// TIA Portal project "1215C_BREAKOUT_BOARD_IO-LINK_TEMPERATURE&TOWERLIGHT" (V19)

(* hardware
DEVICE "BREAKOUT_BOARD_PLC"  S7-1200 Station
   slot 0: "Rack_0"  S7-1200 Rack  Rack  V1.0
   slot 1: "BREAKOUT_BOARD_PLC"  CPU 1215C DC/DC/DC  6ES7 215-1AG40-0XB0  V4.6
DEVICE "BREAKOUT_BOARD_HMI"  KTP400 Basic PN
   slot 0: "BREAKOUT_BOARD_HMI"  KTP400 Basic PN  6AV2 123-2DB03-0AX0  16.0.0.0
   slot 1: "HMI_RT_1"  KTP400 Basic PN  6AV2 123-2DB03-0AX0  16.0.0.0
   slot 5: "BREAKOUT_BOARD_HMI.IE_CP_1"  PROFINET Interface  16.0.0.0
      slot 1: "PROFINET Interface"  PROFINET Interface
         slot 1: "Port_1"  Port
DEVICE "IFM_IO-LINK_MASTER"  GSD.Device.PN
   slot 0: "Rack"  Rack  V1.0
   slot 0: "AL1100"  AL1100  AL1100
      slot 0: "AL1100"  AL1100
      slot 1: "X1"  X1
         slot 1: "Port 1"  Port 1
         slot 2: "Port 2"  Port 2
      slot 1: "4 Ports_1"  4 Ports  AL1100
         slot 0: "IO-Link Master"  IO-Link Master
   slot 1: "IFM ITA2105 IO-Link In  2 Byte + PQI"  IO-Link In  2 Byte + PQI
   slot 2: "Banner TLF100 IO-Link Out 32 Byte + PQI"  IO-Link Out 32 Byte + PQI
   slot 3: "Disabled_P3"  Disabled
   slot 4: "Disabled_P4"  Disabled
DEVICE "SCALANCE XB008"  SCALANCE X-Station
   slot 0: "SCALANCE X rack"  Rail
   slot 0: "8PORT_SWITCH"  6GK5 008-0BA10-1AB2  V1.0
*)

// ===== PLC "BREAKOUT_BOARD_PLC"  CPU 1215C DC/DC/DC =====

VAR_GLOBAL   // PLC tag table "PLC_Outputs"
   "DQ0.0" AT %Q0.0 : Bool;   // Digital Output
   "DQ0.1" AT %Q0.1 : Bool;   // Digital Output
   "DQ0.2" AT %Q0.2 : Bool;   // Digital Output
   "DQ0.3" AT %Q0.3 : Bool;   // Digital Output
   "DQ0.4" AT %Q0.4 : Bool;   // Digital Output
   "DQ0.5" AT %Q0.5 : Bool;   // Digital Output
   "DQ0.6" AT %Q0.6 : Bool;   // Digital Output
   "DQ0.7" AT %Q0.7 : Bool;   // Digital Output
   "DQ1.0" AT %Q1.0 : Bool;   // Digital Output
   "DQ1.1" AT %Q1.1 : Bool;   // Digital Output
   "AQ0.0" AT %QW64 : Word;   // Analog Output
   "AQ0.1" AT %QW66 : Word;   // Analog Output
END_VAR

VAR_GLOBAL   // PLC tag table "PLC_Inputs"
   "DI0.0" AT %I0.0 : Bool;   // Digital Input
   "DI0.1" AT %I0.1 : Bool;   // Digital Input
   "DI0.2" AT %I0.2 : Bool;   // Digital Input
   "DI0.3" AT %I0.3 : Bool;   // Digital Input
   "DI0.4" AT %I0.4 : Bool;   // Digital Input
   "DI0.5" AT %I0.5 : Bool;   // Digital Input
   "DI0.6" AT %I0.6 : Bool;   // Digital Input
   "DI0.7" AT %I0.7 : Bool;   // Digital Input
   "DI1.0" AT %I1.0 : Bool;   // Digital Input
   "DI1.1" AT %I1.1 : Bool;   // Digital Input
   "DI1.2" AT %I1.2 : Bool;   // Digital Input
   "DI1.3" AT %I1.3 : Bool;   // Digital Input
   "DI1.4" AT %I1.4 : Bool;   // Digital Input
   "DI1.5" AT %I1.5 : Bool;   // Digital Input
   "AI0.0" AT %IW64 : Word;   // Analog Input
   "AI0.1" AT %IW66 : Word;   // Analog Input
END_VAR

VAR_GLOBAL   // PLC tag table "System_Tags"
   "Clock_Byte" AT %MB0 : Byte;
   "Clock_10Hz" AT %M0.0 : Bool;
   "Clock_5Hz" AT %M0.1 : Bool;
   "Clock_2.5Hz" AT %M0.2 : Bool;
   "Clock_2Hz" AT %M0.3 : Bool;
   "Clock_1.25Hz" AT %M0.4 : Bool;
   "Clock_1Hz" AT %M0.5 : Bool;
   "Clock_0.625Hz" AT %M0.6 : Bool;
   "Clock_0.5Hz" AT %M0.7 : Bool;
   "System_Byte" AT %MB1 : Byte;
   "FirstScan" AT %M1.0 : Bool;
   "DiagStatusUpdate" AT %M1.1 : Bool;
   "AlwaysTRUE" AT %M1.2 : Bool;
   "AlwaysFALSE" AT %M1.3 : Bool;
END_VAR

VAR_GLOBAL   // PLC tag table "Trigger_Tags"
   "xAQ_Trig" AT %M2.0 : Bool;
   "xTrig2" AT %M2.1 : Bool;
   "xTrig3" AT %M2.2 : Bool;
   "xTrig4" AT %M2.3 : Bool;
   "xTrig5" AT %M2.4 : Bool;
END_VAR

VAR_GLOBAL   // PLC tag table "IO-Link_Tags"
   "IFM_TA2105_Temp" AT %IW68 : Int;   // IO-Link Master X1
   "Banner_TLF100Pro_Byte0" AT %QB2 : Byte;   // IO-Link Master X2
   "Banner_TLF100Pro_Byte1" AT %QB3 : Byte;   // IO-Link Master X2
   "Banner_TLF100Pro_Byte2" AT %QB4 : Byte;   // IO-Link Master X2
   "Banner_TLF100Pro_Byte3" AT %QB5 : Byte;   // IO-Link Master X2
   "Banner_TLF100Pro_Byte4" AT %QB6 : Byte;   // IO-Link Master X2
   "Banner_TLF100Pro_Byte5" AT %QB7 : Byte;   // IO-Link Master X2
   "Banner_TLF100Pro_Byte6" AT %QB8 : Byte;   // IO-Link Master X2
   "Banner_TLF100Pro_Byte7" AT %QB9 : Byte;   // IO-Link Master X2
   "Banner_TLF100Pro_Byte8" AT %QB10 : Byte;   // IO-Link Master X2
   "Banner_TLF100Pro_Byte9" AT %QB11 : Byte;   // IO-Link Master X2
   "Banner_TLF100Pro_Byte10" AT %QB12 : Byte;   // IO-Link Master X2
   "Banner_TLF100Pro_Byte11" AT %QB13 : Byte;   // IO-Link Master X2
   "Banner_TLF100Pro_Byte12" AT %QB14 : Byte;   // IO-Link Master X2
   "Banner_TLF100Pro_Byte13" AT %QB15 : Byte;   // IO-Link Master X2
   "Banner_TLF100Pro_Byte14" AT %QB16 : Byte;   // IO-Link Master X2
   "Banner_TLF100Pro_Byte15" AT %QB17 : Byte;   // IO-Link Master X2
   "Banner_TLF100Pro_Byte16" AT %QB18 : Byte;   // IO-Link Master X2
   "Banner_TLF100Pro_Byte17" AT %QB19 : Byte;   // IO-Link Master X2
   "Banner_TLF100Pro_Byte18" AT %QB20 : Byte;   // IO-Link Master X2
   "Banner_TLF100Pro_Byte19" AT %QB21 : Byte;   // IO-Link Master X2
   "Banner_TLF100Pro_Byte20" AT %QB22 : Byte;   // IO-Link Master X2
   "Banner_TLF100Pro_Byte21" AT %QB23 : Byte;   // IO-Link Master X2
   "Banner_TLF100Pro_Byte22" AT %QB24 : Byte;   // IO-Link Master X2 - Not Used
   "Banner_TLF100Pro_Byte23" AT %QB25 : Byte;   // IO-Link Master X2 - Not Used
   "Banner_TLF100Pro_Byte24" AT %QB26 : Byte;   // IO-Link Master X2 - Not Used
   "Banner_TLF100Pro_Byte25" AT %QB27 : Byte;   // IO-Link Master X2 - Not Used
   "Banner_TLF100Pro_Byte26" AT %QB28 : Byte;   // IO-Link Master X2 - Not Used
   "Banner_TLF100Pro_Byte27" AT %QB29 : Byte;   // IO-Link Master X2 - Not Used
   "Banner_TLF100Pro_Byte28" AT %QB30 : Byte;   // IO-Link Master X2 - Not Used
   "Banner_TLF100Pro_Byte29" AT %QB31 : Byte;   // IO-Link Master X2 - Not Used
   "Banner_TLF100Pro_Byte30" AT %QB32 : Byte;   // IO-Link Master X2 - Not Used
   "Banner_TLF100Pro_Byte31" AT %QB33 : Byte;   // IO-Link Master X2 - Not Used
END_VAR

// folder: WS01_TVET_Workstation/00-I/O_Mapping

DATA_BLOCK "DB001-PLC_I/O"   // DB1
TITLE = PLC I/O Global Database
{ S7_Optimized_Access := 'TRUE' }
VERSION : 0.1
// Variables used to mirror the physical PLC I/O states.
   VAR
      Inputs : Struct   // PLC Inputs Structure
         "xDI0.0" : Bool;
         "xDI0.1" : Bool;
         "xDI0.2" : Bool;
         "xDI0.3" : Bool;
         "xDI0.4" : Bool;
         "xDI0.5" : Bool;
         "xDI0.6" : Bool;
         "xDI0.7" : Bool;
         "xDI1.0" : Bool;
         "xDI1.1" : Bool;
         "xDI1.2" : Bool;
         "xDI1.3" : Bool;
         "xDI1.4" : Bool;
         "xDI1.5" : Bool;
         "rAI0.0_Scaled" : Real;   // 0 to 24648 = 0 to 10 V
         "rAI0.1_Scaled" : Real;   // 0 to 24648 = 0 to 10 V
      END_STRUCT;
      Outputs : Struct   // PLC Outputs Structure
         "xDQ0.0" : Bool;
         "xDQ0.1" : Bool;
         "xDQ0.2" : Bool;
         "xDQ0.3" : Bool;
         "xDQ0.4" : Bool;
         "xDQ0.5" : Bool;
         "xDQ0.6" : Bool;
         "xDQ0.7" : Bool;
         "xDQ1.0" : Bool;
         "xDQ1.1" : Bool;
         "iAQ0.0_RAW" : Int := 0;
         "rAQ0.0_Scaled" : Real;   // 0 to 24648 = 0 to 20 mA
         "iAQ0.1_RAW" : Int := 0;
         "rAQ0.1_Scaled" : Real;   // 0 to 24648 = 0 to 20 mA
      END_STRUCT;
   END_VAR
BEGIN
END_DATA_BLOCK

DATA_BLOCK "DB003-IO-Link_I/O"   // DB3
TITLE = IO-Link I/O Global Database
{ S7_Optimized_Access := 'TRUE' }
VERSION : 0.1
// Variables used to mirror the physical IO-Link I/O states.
   VAR
      Inputs : Struct   // IO-Link Inputs Structure
         wTemp_RAW : Word;   // Temperature Sensor Scaled Value
      END_STRUCT;
      Outputs : Struct   // IO-Link Outputs Structure
         TL_Byte_Array : Array[0..21] of Byte;   // Tower Light Byte Array
      END_STRUCT;
   END_VAR
BEGIN
END_DATA_BLOCK

// folder: WS01_TVET_Workstation/01-DateTime

DATA_BLOCK "DB002-DateTime"   // DB2
TITLE = PLC Date/Time Global Database
{ S7_Optimized_Access := 'TRUE' }
VERSION : 0.1
// Variables used to store the PLC date/time & custom date/time formatting.
   VAR
      RD_LOC_T_Ret : Int := 0;   // Return value for Read Local Time Block
      LOCAL_DTL : DTL := DTL#1970-01-01-00:00:00;   // RAW DTL
      "Date" : Date := D#1990-01-01;   // RAW Date
      "Time" : Time_Of_Day := TOD#00:00:00;   // RAW Time
      DTLtoString_Ret : String;   // Return value for DTL to String Block
      sCustomDate_YY : String := '';   // Custom year
      sCustomDate_MM : String := '';   // Custom month
      sCustomDate_DD : String := '';   // Custom Day
      sCustomTime_HH : String := '';   // Custom hour
      sCustomTime_MM : String := '';   // Custom minute
      sCustomDate_DDMMYY : String := '';   // Custom date format
      sCustomTime_HHMM : String := '';   // Custom time format
   END_VAR
BEGIN
END_DATA_BLOCK

// folder: WS01_TVET_Workstation/02-IOLink_Control

DATA_BLOCK "DB003-IOLink_Data"   // DB4
TITLE = IO-Link Data Global Database
{ S7_Optimized_Access := 'TRUE' }
VERSION : 0.1
// Variables used to process data from connected devices.
   VAR
      TempSensor_Data : Struct   // Temperature Sensor Data Structure
         rDeg_C : Real;   // Degrees Celsius
         rDeg_F : Real;   // Degrees Fahrenheit
      END_STRUCT;
      TL_ProcessData : Struct   // Tower Light Process Data Structure
         Animations : Struct   // Animation Parameters Structure
            iOff : Int := 0;   // Animations
            iSteady : Int := 1;   // Animations
            iFlash : Int := 2;   // Animations
            i2ColourFlash : Int := 3;   // Animations
            i2ColourShift : Int := 4;   // Animations
            iEndsSteady : Int := 5;   // Animations
            iEndsFlash : Int := 6;   // Animations
            iScroll : Int := 7;   // Animations
            iCenterScroll : Int := 8;   // Animations
            iBounce : Int := 9;   // Animations
            iCenterBounce : Int := 10;   // Animations
            iIntensitySweep : Int := 11;   // Animations
            i2ColourSweep : Int := 12;   // Animations
            iSpectrum : Int := 13;   // Animations
            iLevelSteady : Int := 14;   // Animations
            iLevelFlash : Int := 15;   // Animations
         END_STRUCT;
         Colours : Struct   // Colour Parameters Structure
            iGreen : Int := 0;   // Colours
            iRed : Int := 1;   // Colours
            iOrange : Int := 2;   // Colours
            iAmber : Int := 3;   // Colours
            iYellow : Int := 4;   // Colours
            iLimeGreen : Int := 5;   // Colours
            iSpringGreen : Int := 6;   // Colours
            iCyan : Int := 7;   // Colours
            iSkyBlue : Int := 8;   // Colours
            iBlue : Int := 9;   // Colours
            iViolet : Int := 10;   // Colours
            iMegenta : Int := 11;   // Colours
            iRose : Int := 12;   // Colours
            iDaylightWhite : Int := 13;   // Colours
         END_STRUCT;
         ColourIntensities : Struct   // Colour Intensity Parameters Structure
            iHigh : Int := 0;   // Colour Intensity
            iLow : Int := 1;   // Colour Intensity
            iMedium : Int := 2;   // Colour Intensity
            iOff : Int := 3;   // Colour Intensity
         END_STRUCT;
         Speeds : Struct   // Speed Parameters Structure
            iMedium : Int := 0;   // Speed
            iFast : Int := 1;   // Speed
            iSlow : Int := 2;   // Speed
         END_STRUCT;
         PulsePatterns : Struct   // Pulse Pattern Parameters Structure
            iNormal : Int := 0;   // Pulse Pattern
            iStrobe : Int := 1;   // Pulse Pattern
            i3Pulse : Int := 2;   // Pulse Pattern
            iSOS : Int := 3;   // Pulse Pattern
            iRandom : Int := 4;   // Pulse Pattern
         END_STRUCT;
         ScrollStyles : Struct   // Scroll Style Parameters Structure
            iSolid : Int := 0;   // Scroll Style
            iTail : Int := 1;   // Scroll Style
            iRipple : Int := 2;   // Scroll Style
         END_STRUCT;
         Directions : Struct   // Direction Parameters Structure
            xUp : Bool := FALSE;   // Direction
            xDown : Bool := TRUE;   // Direction
         END_STRUCT;
         iColourWidthPercent : Int := 100;   // Percent Width of Colour (1-100)
         AudibleTypes : Struct   // Audible Type Parameters Structure
            iPulse : Int := 0;   // Audible Type
            iWobble : Int := 1;   // Audible Type
            iStrobe : Int := 2;   // Audible Type
            iWhoop : Int := 4;   // Audible Type
            iStaccato : Int := 5;   // Audible Type
            iSiren : Int := 6;   // Audible Type
            iContinuous1 : Int := 8;   // Audible Type
            iContinuous2 : Int := 9;   // Audible Type
            iJungle : Int := 16;   // Audible Type
            iMelody1 : Int := 17;   // Audible Type
            iMelody2 : Int := 18;   // Audible Type
            iMelody3 : Int := 19;   // Audible Type
         END_STRUCT;
         AudibleVolumes : Struct   // Audible Volume Parameters Structure
            iOff : Int := 0;   // Audible Volume
            iLow : Int := 1;   // Audible Volume
            iMedium : Int := 2;   // Audible Volume
            iHigh : Int := 3;   // Audible Volume
         END_STRUCT;
      END_STRUCT;
   END_VAR
BEGIN
END_DATA_BLOCK

// folder: WS01_TVET_Workstation/03-HMI_Control

DATA_BLOCK "DB005-HMI_Data"   // DB5
TITLE = HMI Data Global Database
{ S7_Optimized_Access := 'TRUE' }
VERSION : 0.1
// Variables used to process data from the HMI.
   VAR
      iScreen_Number : UInt;   // HMI Active Screen Number
      TowerLight : Struct   // Tower Light HMI Variables Structure
         Segment1 : Struct   // Segment 1 Structure
            iAnimate : Int;   // Animations
            iSavedAnimate : Int;   // Saved Animation Value
            iColour1 : Int;   // Colour1 Colours
            iColour2 : Int;   // Colour2 Colours
            iSpeed : Int;   // Speeds
            "iClrWidth%" : Int := 100;   // Colour Width Percentage
         END_STRUCT;
         Segment2 : Struct   // Segment 2 Structure
            iAnimate : Int;   // Animations
            iSavedAnimate : Int;   // Saved Animation Value
            iColour1 : Int;   // Colour1 Colours
            iColour2 : Int;   // Colour2 Colours
            iSpeed : Int;   // Speeds
            "iClrWidth%" : Int := 100;   // Colour Width Percentage
         END_STRUCT;
         Segment3 : Struct   // Segment 3 Structure
            iAnimate : Int;   // Animations
            iSavedAnimate : Int;   // Saved Animation Value
            iColour1 : Int;   // Colour1 Colours
            iColour2 : Int;   // Colour2 Colours
            iSpeed : Int;   // Speeds
            "iClrWidth%" : Int := 100;   // Colour Width Percentage
         END_STRUCT;
         Audible : Struct   // Audible (Sound) Structure
            iType : Int;   // Types
            iVolume : Int;   // Volumes
            iSavedVolume : Int;   // Saved Volume Value
         END_STRUCT;
         xSave_Config : Bool;   // Save Tower Light Configs Button
      END_STRUCT;
   END_VAR
BEGIN
END_DATA_BLOCK

// folder: (top level)

ORGANIZATION_BLOCK "Main"   // OB1, LAD, ProgramCycle
TITLE = "Main Program Sweep (Cycle)"
{ S7_Optimized_Access := 'TRUE' }
VERSION : 0.1
   VAR_INPUT
      Initial_Call : Bool;   // Initial call of this OB
      Remanence : Bool;   // =True, if remanent data are available
   END_VAR
BEGIN

REGION Network 1 (SCL): ================= PROGRAM_INFORMATION =================
   (*
   ==================================================================
   ********************* PLC I/O BREAKOUT BOARD *********************
   ==================================================================

   TVET Workstation WS01:
   1215C DC/DC/DC - 6ES7215-1AG40-0XB0 - IP: 192.168.0.175/24

   KTP400 HMI - 6AV2123-2DB03-0AX0 - IP: 192.168.0.176/24

   IFM IO-Link Master - AL1100 - IP: 192.168.0.177/24

   =======================================================================

   The program has 4 main sections:
   - Date/Time Handler,
   - I/O Handlers,
   - IO-Link Devices Handler,
   - HMI Handler.

   Date/Time Handler FC:
   - local PLC date/time is read & formatted into a 24HR time & DD/MM/YYYY.

   I/O Handler FCs:
   - maps the physical PLC inputs & outputs to corresponding tags in DB001,
   - handles scaling of the PLC Analog I/O,
   - maps the IO-Link inputs & outputs to corresponding tags in DB003,
   - ensures that physical I/O tags are only used once in the code.

   IO-Link Device Handler FCs:
   - connected IO-Link devices are controlled in this section:
       - the temperature sensor conversion logic is handled by an IFM
         provided FC which scales the input value & converts to Fahrenheit.
       - the tower light ON/OFF logic is handled by the TowerLight Handler FC.
   - create & call new FC's for any additional IO-Link devices that may
     get added.

   Additional Notes:
   PLC Tags grouped according to their use/function.

   =======================================================================

   Analog Input Technical data:
   - Number of inputs: 2
   - Type: Voltage (single-ended)
   - Full-scale range: 0 to 10 V
   - Full-scale range (data word): 0 to 27648
   - Overshoot range: 10.001 to 11.759 V
   - Overshoot range (data word): 27649 to 32511
   - Overflow range: 11.760 to 11.852 V
   - Overflow range (data word): 32512 to 32767
   - Resolution: 10 bits
   - Maximum withstand voltage: 35 V DC
   - Smoothing: None, Weak, Medium, or Strong
   - Noise rejection: 10, 50, or 60 Hz
   - Impedance: ≥100 KΩ
   - Isolation (field side to logic): None
   - Accuracy (25 °C / -20 to 60 °C): 3.0% / 3.5% of full-scale
   - Cable length (meters): 100 m, shielded twisted pair
   - Rated range: 0     = 0 V
                  34    = 12 mV
                  20736 = 7.5 V
                  27648 = 10 V

   =======================================================================

   Analog Output Technical data:
   - Number of outputs: 2
   - Type: Current
   - Full-scale range: 0 to 20 mA
   - Full-scale range (data word): 0 to 27648
   - Overshoot range: 20.01 to 23.52 mA
   - Overshoot range (data word): 27649 to 32511
   - Overflow range data word: 32512 to 32767
   - Resolution: 10 bits
   - Output drive impedance: ≤500 Ω max
   - Isolation (field side to logic): None
   - Accuracy (25 °C / -20 to 60 °C): 3.0% / 3.5% of full-scale
   - Settling time: 2 ms
   - Cable length (meters): 100 m, shielded twisted pair
   - Rated range: 0     = 0 mA
                  34    = 0.0247 mA
                  20736 = 15 mA
                  27648 = 20 mA

   =======================================================================

   TA2105 IO-Link Temperature Transmitter documentation:
   https://www.ifm.com/us/en/product/TA2105#documents

   Process Data In length = 2bytes

   The IO-Link Inputs screen on the HMI displays a bar graph of the current
   measured temperature for the sensor connected to port X1.

   =======================================================================

   TLF100Pro IO-Link Tower Light Data Reference Guide:
   www.bannerengineering.com/us/en/products/part.812293.html

   Process Data Out length = 22bytes

   Modes:
   - Segment Mode
   - Run Mode
   - Advanced Mode
   - Level Mode

   We will be using the "Advanced Mode" to configure Segments 1, 2, 3
   and Audible. Segment 4 can be ignored as it is not applicable to
   this tower light model.

   The function interface contains a list of the available parameters
   that can be used to set segment bytes.

   Each colour segment has 5 bytes that need to be set with a
   corresponding constant value to configure the segment.

   The audible (segment) has 2 bytes that need to be set with a
   corresponding constant value.

   Segment bytes are defined as follows:
   -----------------------------
   > Segement 1 - byte 21 to 17:
       - 21 = Animation (8bits)
       - 20 = Colour1 (5bits) + Intensity (3bits)
       - 19 = Colour2 (5bits) + Intensity (3bits)
       - 18 = Speed (2bits) + Pulse Pattern (3bits) + Style (2bits) + Direction (1bit)
       - 17 = Colour Width Percentage (1-100)
   -----------------------------
   > Segement 2 - byte 16 to 12:
       - 16 = Animation (8bits)
       - 15 = Colour1 (5bits) + Intensity (3bits)
       - 14 = Colour2 (5bits) + Intensity (3bits)
       - 13 = Speed (2bits) + Pulse Pattern (3bits) + Style (2bits) + Direction (1bit)
       - 12 = Colour Width Percentage (1-100)
   ----------------------------
   > Segement 3 - byte 11 to 7:
       - 11 = Animation (8bits)
       - 10 = Colour1 (5bits) + Intensity (3bits)
       - 09 = Colour2 (5bits) + Intensity (3bits)
       - 08 = Speed (2bits) + Pulse Pattern (3bits) + Style (2bits) + Direction (1bit)
       - 07 = Colour Width Percentage (1-100)
   ---------------------------
   > Segement 4 - byte 6 to 2: !!NOT USED!!
       - 06 = Animation (8bits)
       - 05 = Colour1 (5bits) + Intensity (3bits)
       - 04 = Colour2 (5bits) + Intensity (3bits)
       - 03 = Speed (2bits) + Pulse Pattern (3bits) + Style (2bits) + Direction (1bit)
       - 02 = Colour Width Percentage (1-100)
   ------------------------
   > Audible - byte 1 to 0:
       - 01 = Type (8bits)
       - 00 = Volume (8bits)

   Some segment bytes are divided into sub-indexes depending on the 
   functions available for a particular byte.

   Since we are aiming at creating basic functionality
   (basic solid or flashing colours & sound)
   we will ignore many of the sub-indexes functions & simply set the
   entire byte with a single parameter constant.

   Segment parameters are set via the HMI and controlled via input
   switches.

   =======================================================================
   *)
END_REGION

REGION Network 2: ================= LOCAL_DATE/TIME =================
END_REGION

REGION Network 3: Call the Date/Time Handler Function
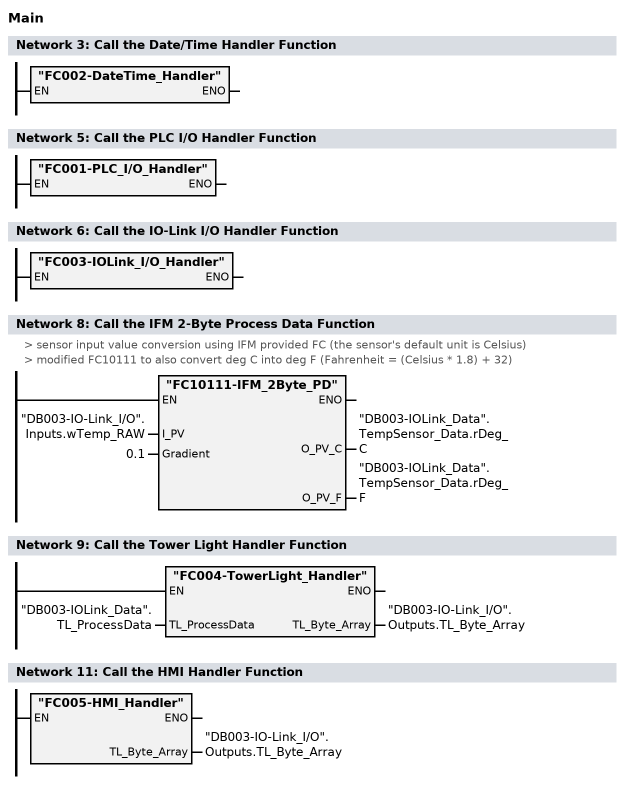
   RUNG wire#powerrail
      "FC002-DateTime_Handler"()
   END_RUNG
   // the same network as SCL:
   "FC002-DateTime_Handler"();
END_REGION

REGION Network 4: ================= I/O_MAPPING =================
END_REGION

REGION Network 5: Call the PLC I/O Handler Function
   RUNG wire#powerrail
      "FC001-PLC_I/O_Handler"()
   END_RUNG
   // the same network as SCL:
   "FC001-PLC_I/O_Handler"();
END_REGION

REGION Network 6: Call the IO-Link I/O Handler Function
   RUNG wire#powerrail
      "FC003-IOLink_I/O_Handler"()
   END_RUNG
   // the same network as SCL:
   "FC003-IOLink_I/O_Handler"();
END_REGION

REGION Network 7: ================= IO-LINK_DEVICES =================
END_REGION

REGION Network 8: Call the IFM 2-Byte Process Data Function
   // > sensor input value conversion using IFM provided FC (the sensor's default unit is Celsius)
   // > modified FC10111 to also convert deg C into deg F (Fahrenheit = (Celsius * 1.8) + 32)
   RUNG wire#powerrail
      "FC10111-IFM_2Byte_PD"(I_PV := "DB003-IO-Link_I/O".Inputs.wTemp_RAW, Gradient := 0.1, O_PV_C => "DB003-IOLink_Data".TempSensor_Data.rDeg_C, O_PV_F => "DB003-IOLink_Data".TempSensor_Data.rDeg_F)
   END_RUNG
   // the same network as SCL:
   "FC10111-IFM_2Byte_PD"(I_PV := "DB003-IO-Link_I/O".Inputs.wTemp_RAW,
                          Gradient := 0.1,
                          O_PV_C => "DB003-IOLink_Data".TempSensor_Data.rDeg_C,
                          O_PV_F => "DB003-IOLink_Data".TempSensor_Data.rDeg_F);
END_REGION

REGION Network 9: Call the Tower Light Handler Function
   RUNG wire#powerrail
      "FC004-TowerLight_Handler"(TL_ProcessData := "DB003-IOLink_Data".TL_ProcessData, TL_Byte_Array => "DB003-IO-Link_I/O".Outputs.TL_Byte_Array)
   END_RUNG
   // the same network as SCL:
   "FC004-TowerLight_Handler"(TL_ProcessData := "DB003-IOLink_Data".TL_ProcessData,
                           TL_Byte_Array => "DB003-IO-Link_I/O".Outputs.TL_Byte_Array);
END_REGION

REGION Network 10: ================= HMI_CONTROL =================
END_REGION

REGION Network 11: Call the HMI Handler Function
   RUNG wire#powerrail
      "FC005-HMI_Handler"(TL_Byte_Array => "DB003-IO-Link_I/O".Outputs.TL_Byte_Array)
   END_RUNG
   // the same network as SCL:
   "FC005-HMI_Handler"(TL_Byte_Array => "DB003-IO-Link_I/O".Outputs.TL_Byte_Array);
END_REGION
END_ORGANIZATION_BLOCK

// folder: WS01_TVET_Workstation/00-I/O_Mapping

FUNCTION "FC001-PLC_I/O_Handler" : Void   // FC1, LAD
TITLE = PLC Input Output Handler
{ S7_Optimized_Access := 'TRUE' }
VERSION : 0.1
// This function block is for interfacing the physical PLC input/output connections to a Global DB's (DB001-PLC_I/O for ).
   VAR_TEMP
      "rAI0.0_Temp" : Real;
      "rAI0.1_Temp" : Real;
      "rAQ0.0_Temp" : Real;
      "rAQ0.1_Temp" : Real;
   END_VAR
   VAR_TEMP   // added for the SCL form of the ladder/FBD networks
      _w1 : Bool;
   END_VAR
BEGIN

REGION Network 1: ================= DIGITAL_INPUTS =================
END_REGION

REGION Network 2: BANK_0
   // > DI0.0 - DI0.7
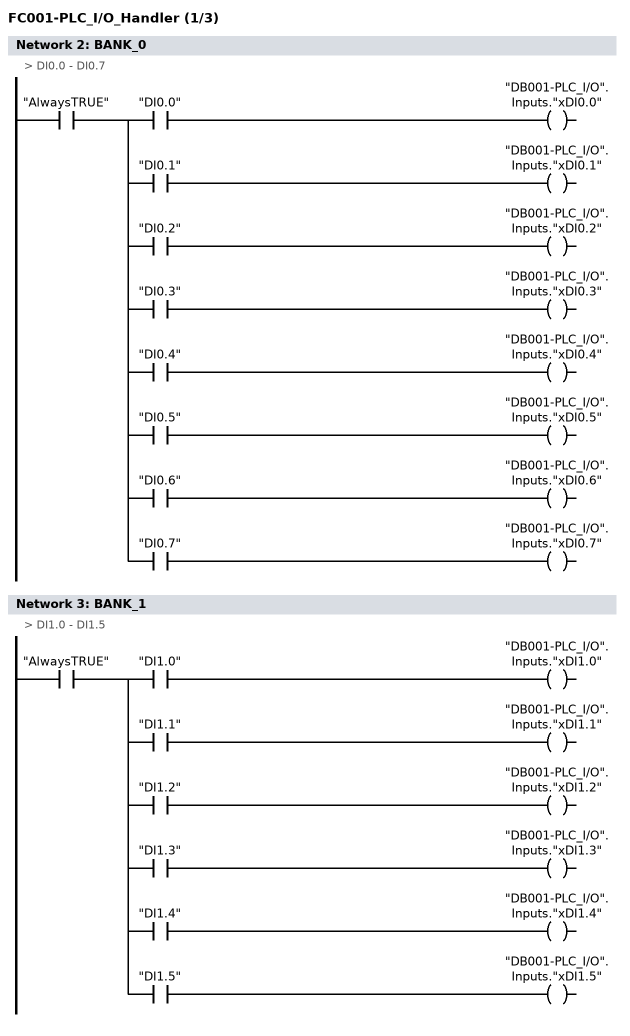
   RUNG wire#powerrail
      Contact( "AlwaysTRUE" )
      wire#w1
      Contact( "DI0.0" )
      Coil( "DB001-PLC_I/O".Inputs."xDI0.0" )
   END_RUNG
   RUNG wire#w1
      Contact( "DI0.1" )
      Coil( "DB001-PLC_I/O".Inputs."xDI0.1" )
   END_RUNG
   RUNG wire#w1
      Contact( "DI0.2" )
      Coil( "DB001-PLC_I/O".Inputs."xDI0.2" )
   END_RUNG
   RUNG wire#w1
      Contact( "DI0.3" )
      Coil( "DB001-PLC_I/O".Inputs."xDI0.3" )
   END_RUNG
   RUNG wire#w1
      Contact( "DI0.4" )
      Coil( "DB001-PLC_I/O".Inputs."xDI0.4" )
   END_RUNG
   RUNG wire#w1
      Contact( "DI0.5" )
      Coil( "DB001-PLC_I/O".Inputs."xDI0.5" )
   END_RUNG
   RUNG wire#w1
      Contact( "DI0.6" )
      Coil( "DB001-PLC_I/O".Inputs."xDI0.6" )
   END_RUNG
   RUNG wire#w1
      Contact( "DI0.7" )
      Coil( "DB001-PLC_I/O".Inputs."xDI0.7" )
   END_RUNG
   // the same network as SCL:
   "DB001-PLC_I/O".Inputs."xDI0.0" := "AlwaysTRUE" AND "DI0.0";
   "DB001-PLC_I/O".Inputs."xDI0.1" := "AlwaysTRUE" AND "DI0.1";
   "DB001-PLC_I/O".Inputs."xDI0.2" := "AlwaysTRUE" AND "DI0.2";
   "DB001-PLC_I/O".Inputs."xDI0.3" := "AlwaysTRUE" AND "DI0.3";
   "DB001-PLC_I/O".Inputs."xDI0.4" := "AlwaysTRUE" AND "DI0.4";
   "DB001-PLC_I/O".Inputs."xDI0.5" := "AlwaysTRUE" AND "DI0.5";
   "DB001-PLC_I/O".Inputs."xDI0.6" := "AlwaysTRUE" AND "DI0.6";
   "DB001-PLC_I/O".Inputs."xDI0.7" := "AlwaysTRUE" AND "DI0.7";
END_REGION

REGION Network 3: BANK_1
   // > DI1.0 - DI1.5
   RUNG wire#powerrail
      Contact( "AlwaysTRUE" )
      wire#w1
      Contact( "DI1.0" )
      Coil( "DB001-PLC_I/O".Inputs."xDI1.0" )
   END_RUNG
   RUNG wire#w1
      Contact( "DI1.1" )
      Coil( "DB001-PLC_I/O".Inputs."xDI1.1" )
   END_RUNG
   RUNG wire#w1
      Contact( "DI1.2" )
      Coil( "DB001-PLC_I/O".Inputs."xDI1.2" )
   END_RUNG
   RUNG wire#w1
      Contact( "DI1.3" )
      Coil( "DB001-PLC_I/O".Inputs."xDI1.3" )
   END_RUNG
   RUNG wire#w1
      Contact( "DI1.4" )
      Coil( "DB001-PLC_I/O".Inputs."xDI1.4" )
   END_RUNG
   RUNG wire#w1
      Contact( "DI1.5" )
      Coil( "DB001-PLC_I/O".Inputs."xDI1.5" )
   END_RUNG
   // the same network as SCL:
   "DB001-PLC_I/O".Inputs."xDI1.0" := "AlwaysTRUE" AND "DI1.0";
   "DB001-PLC_I/O".Inputs."xDI1.1" := "AlwaysTRUE" AND "DI1.1";
   "DB001-PLC_I/O".Inputs."xDI1.2" := "AlwaysTRUE" AND "DI1.2";
   "DB001-PLC_I/O".Inputs."xDI1.3" := "AlwaysTRUE" AND "DI1.3";
   "DB001-PLC_I/O".Inputs."xDI1.4" := "AlwaysTRUE" AND "DI1.4";
   "DB001-PLC_I/O".Inputs."xDI1.5" := "AlwaysTRUE" AND "DI1.5";
END_REGION

REGION Network 4: ================= DIGITAL_OUTPUTS =================
END_REGION

REGION Network 5: BANK_0
   // > DQ0.0 - DQ0.7
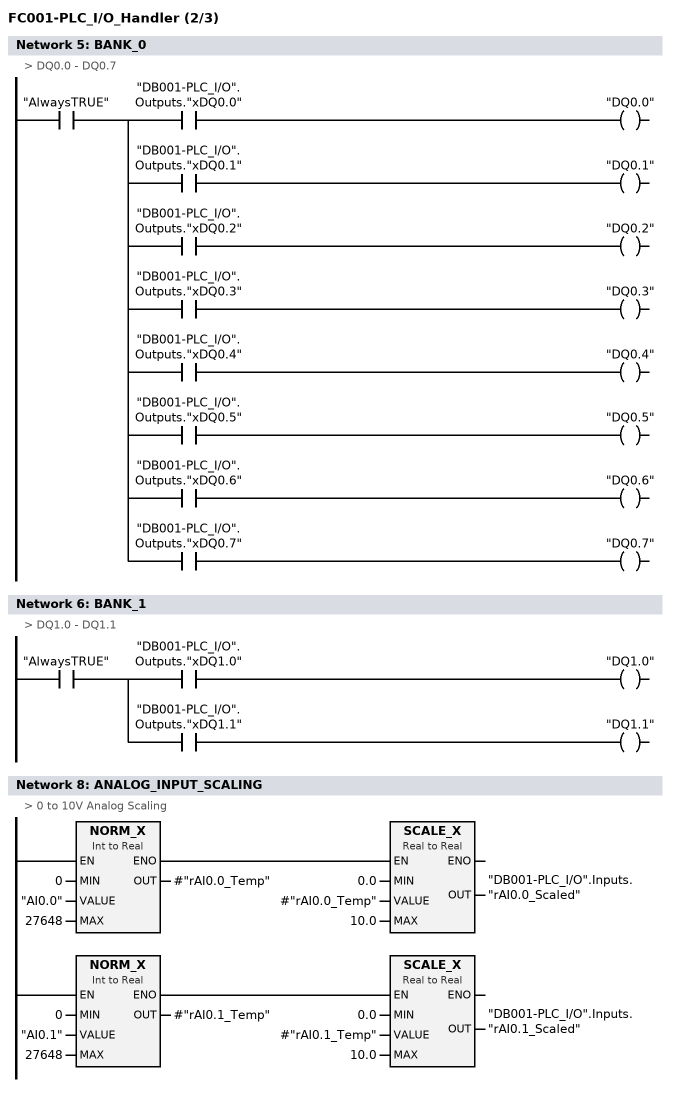
   RUNG wire#powerrail
      Contact( "AlwaysTRUE" )
      wire#w1
      Contact( "DB001-PLC_I/O".Outputs."xDQ0.0" )
      Coil( "DQ0.0" )
   END_RUNG
   RUNG wire#w1
      Contact( "DB001-PLC_I/O".Outputs."xDQ0.1" )
      Coil( "DQ0.1" )
   END_RUNG
   RUNG wire#w1
      Contact( "DB001-PLC_I/O".Outputs."xDQ0.2" )
      Coil( "DQ0.2" )
   END_RUNG
   RUNG wire#w1
      Contact( "DB001-PLC_I/O".Outputs."xDQ0.3" )
      Coil( "DQ0.3" )
   END_RUNG
   RUNG wire#w1
      Contact( "DB001-PLC_I/O".Outputs."xDQ0.4" )
      Coil( "DQ0.4" )
   END_RUNG
   RUNG wire#w1
      Contact( "DB001-PLC_I/O".Outputs."xDQ0.5" )
      Coil( "DQ0.5" )
   END_RUNG
   RUNG wire#w1
      Contact( "DB001-PLC_I/O".Outputs."xDQ0.6" )
      Coil( "DQ0.6" )
   END_RUNG
   RUNG wire#w1
      Contact( "DB001-PLC_I/O".Outputs."xDQ0.7" )
      Coil( "DQ0.7" )
   END_RUNG
   // the same network as SCL:
   "DQ0.0" := "AlwaysTRUE" AND "DB001-PLC_I/O".Outputs."xDQ0.0";
   "DQ0.1" := "AlwaysTRUE" AND "DB001-PLC_I/O".Outputs."xDQ0.1";
   "DQ0.2" := "AlwaysTRUE" AND "DB001-PLC_I/O".Outputs."xDQ0.2";
   "DQ0.3" := "AlwaysTRUE" AND "DB001-PLC_I/O".Outputs."xDQ0.3";
   "DQ0.4" := "AlwaysTRUE" AND "DB001-PLC_I/O".Outputs."xDQ0.4";
   "DQ0.5" := "AlwaysTRUE" AND "DB001-PLC_I/O".Outputs."xDQ0.5";
   "DQ0.6" := "AlwaysTRUE" AND "DB001-PLC_I/O".Outputs."xDQ0.6";
   "DQ0.7" := "AlwaysTRUE" AND "DB001-PLC_I/O".Outputs."xDQ0.7";
END_REGION

REGION Network 6: BANK_1
   // > DQ1.0 - DQ1.1
   RUNG wire#powerrail
      Contact( "AlwaysTRUE" )
      wire#w1
      Contact( "DB001-PLC_I/O".Outputs."xDQ1.0" )
      Coil( "DQ1.0" )
   END_RUNG
   RUNG wire#w1
      Contact( "DB001-PLC_I/O".Outputs."xDQ1.1" )
      Coil( "DQ1.1" )
   END_RUNG
   // the same network as SCL:
   "DQ1.0" := "AlwaysTRUE" AND "DB001-PLC_I/O".Outputs."xDQ1.0";
   "DQ1.1" := "AlwaysTRUE" AND "DB001-PLC_I/O".Outputs."xDQ1.1";
END_REGION

REGION Network 7: ================= ANALOG_PROCESSING =================
END_REGION

REGION Network 8: ANALOG_INPUT_SCALING
   // > 0 to 10V Analog Scaling
   RUNG wire#powerrail
      { S7_Templates := "[SrcType := Int, DestType := Real]" } Normalize(min := 0, value := "AI0.0", max := 27648, out => #"rAI0.0_Temp")
      { S7_Templates := "[SrcType := Real, DestType := Real]" } Scale(min := 0.0, value := #"rAI0.0_Temp", max := 10.0, out => "DB001-PLC_I/O".Inputs."rAI0.0_Scaled")
   END_RUNG
   RUNG wire#powerrail
      { S7_Templates := "[SrcType := Int, DestType := Real]" } Normalize(min := 0, value := "AI0.1", max := 27648, out => #"rAI0.1_Temp")
      { S7_Templates := "[SrcType := Real, DestType := Real]" } Scale(min := 0.0, value := #"rAI0.1_Temp", max := 10.0, out => "DB001-PLC_I/O".Inputs."rAI0.1_Scaled")
   END_RUNG
   // the same network as SCL:
   #"rAI0.0_Temp" := NORM_X(MIN := 0, VALUE := "AI0.0", MAX := 27648);
   "DB001-PLC_I/O".Inputs."rAI0.0_Scaled" := SCALE_X(MIN := 0.0, VALUE := #"rAI0.0_Temp", MAX := 10.0);
   #"rAI0.1_Temp" := NORM_X(MIN := 0, VALUE := "AI0.1", MAX := 27648);
   "DB001-PLC_I/O".Inputs."rAI0.1_Scaled" := SCALE_X(MIN := 0.0, VALUE := #"rAI0.1_Temp", MAX := 10.0);
END_REGION

REGION Network 9: ANALOG_OUTPUT_SCALING
   // > 0 to 20mA Analog Scaling
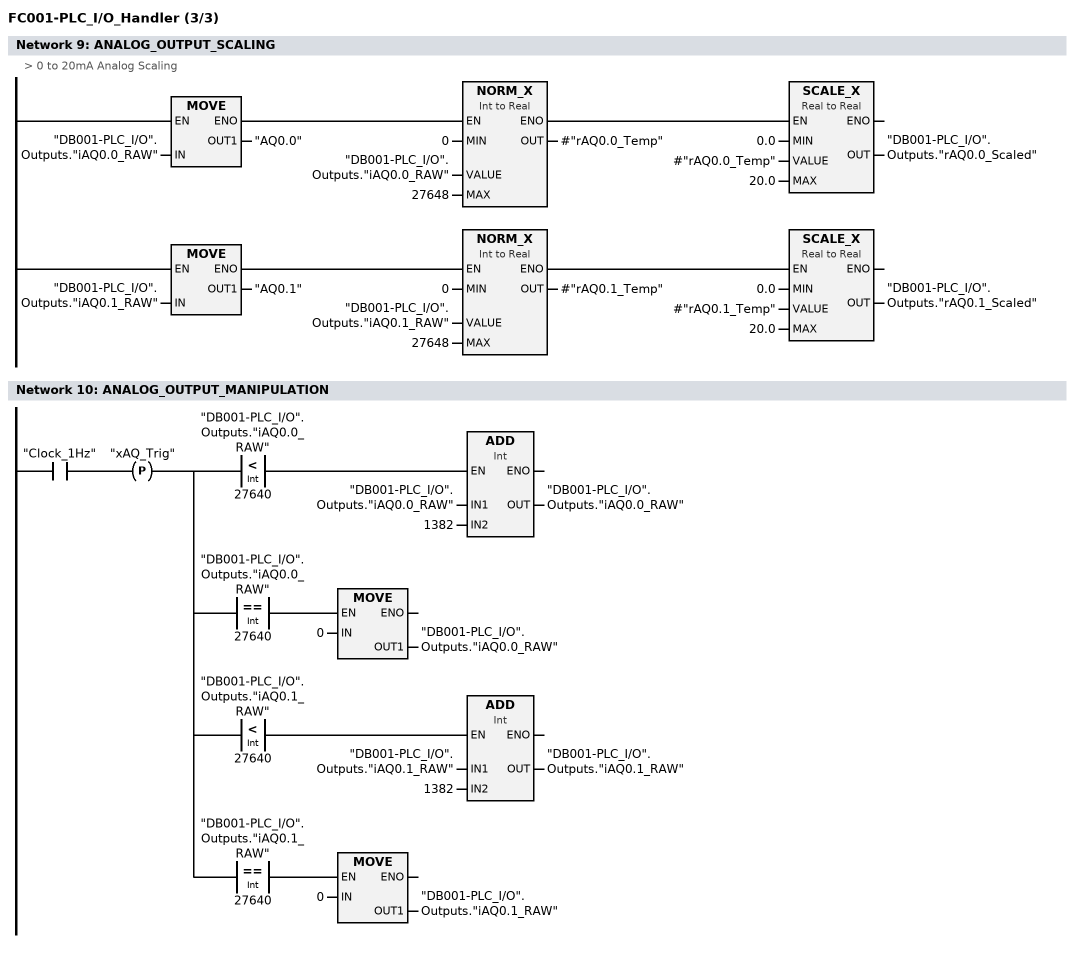
   RUNG wire#powerrail
      Move(in := "DB001-PLC_I/O".Outputs."iAQ0.0_RAW", out1 => "AQ0.0")
      { S7_Templates := "[SrcType := Int, DestType := Real]" } Normalize(min := 0, value := "DB001-PLC_I/O".Outputs."iAQ0.0_RAW", max := 27648, out => #"rAQ0.0_Temp")
      { S7_Templates := "[SrcType := Real, DestType := Real]" } Scale(min := 0.0, value := #"rAQ0.0_Temp", max := 20.0, out => "DB001-PLC_I/O".Outputs."rAQ0.0_Scaled")
   END_RUNG
   RUNG wire#powerrail
      Move(in := "DB001-PLC_I/O".Outputs."iAQ0.1_RAW", out1 => "AQ0.1")
      { S7_Templates := "[SrcType := Int, DestType := Real]" } Normalize(min := 0, value := "DB001-PLC_I/O".Outputs."iAQ0.1_RAW", max := 27648, out => #"rAQ0.1_Temp")
      { S7_Templates := "[SrcType := Real, DestType := Real]" } Scale(min := 0.0, value := #"rAQ0.1_Temp", max := 20.0, out => "DB001-PLC_I/O".Outputs."rAQ0.1_Scaled")
   END_RUNG
   // the same network as SCL:
   "AQ0.0" := "DB001-PLC_I/O".Outputs."iAQ0.0_RAW";
   #"rAQ0.0_Temp" := NORM_X(MIN := 0, VALUE := "DB001-PLC_I/O".Outputs."iAQ0.0_RAW", MAX := 27648);
   "DB001-PLC_I/O".Outputs."rAQ0.0_Scaled" := SCALE_X(MIN := 0.0, VALUE := #"rAQ0.0_Temp", MAX := 20.0);
   "AQ0.1" := "DB001-PLC_I/O".Outputs."iAQ0.1_RAW";
   #"rAQ0.1_Temp" := NORM_X(MIN := 0, VALUE := "DB001-PLC_I/O".Outputs."iAQ0.1_RAW", MAX := 27648);
   "DB001-PLC_I/O".Outputs."rAQ0.1_Scaled" := SCALE_X(MIN := 0.0, VALUE := #"rAQ0.1_Temp", MAX := 20.0);
END_REGION
